// TIA Portal project "SMSS-ENLAB-01-003-1508-012-PLC-B_V13_SP1_1_V17" (V17)

(* hardware
DEVICE "SIMATIC 1200 station_1"  S71200.Device
   slot 0: "S7-1200 rack"  Rack  V1.0
   slot 1: "S7-1200"  CPU 1214C DC/DC/DC  6ES7 214-1AG40-0XB0  V4.5
   slot 2: "DI16 x 24VDC_1"  6ES7 221-1BH30-0XB0  V1.0
   slot 3: "DI8 x 24VDC_1"  6ES7 221-1BF30-0XB0  V1.0
   slot 4: "DQ16 x 24VDC_1"  6ES7 222-1BH30-0XB0  V1.0
DEVICE "HMI"  KTP600 Basic mono PN
   slot 0: "HMI"  HMI  6AV6 647-0AB11-3AX0  12.0.0.0
   slot 1: "HMI_RT_1"  KTP600 Basic mono PN  6AV6 647-0AB11-3AX0  12.0.0.0
   slot 5: "IE_CP_1"  PROFINET Interface  IE_CP  V7.1.0
      slot 1: "PROFINET_Interface_1"  PROFINET Interface
         slot 1: "PORT_1"  Port  1.0.0.0
DEVICE "ET 200S station_1"  ET 200S station
   slot 0: "Rack"  Rail
   slot 0: "IO device_1"  IM 151-3 PN ST  6ES7 151-3AA23-0AB0  V7.0
   slot 1: "PM-E 24VDC_1"  PM-E 24VDC  6ES7 138-4CA01-0AA0
   slot 2: "8DI x 24VDC_1"  8DI DC24V  6ES7 131-4BF00-0AA0
   slot 3: "8DI x 24VDC / SRC ST_1"  8DI DC24V/SRC ST  6ES7 131-4BF50-0AA0
   slot 4: "8DO x 24VDC / 0.5A_1"  8DO DC24V/0.5A  6ES7 132-4BF00-0AA0
DEVICE "CSM"  SCALANCE X-Station
   slot 0: "SCALANCE X rack"  Rail
   slot 0: "CSM 1277 Simatic Net"  6GK7 277-1AA10-0AA0  V1.0
*)

// ===== PLC "S7-1200"  CPU 1214C DC/DC/DC =====

VAR_GLOBAL   // PLC tag table "Default tag table"
   "Flag Negatif Imaje Not ready" AT %M500.2 : Bool;
   "RSAddReject1" AT %I5.5 : Bool;
   "Flag Modu Motor" AT %M300.0 : Bool;
   "RSAddReject2" AT %I5.6 : Bool;
   "PneuAddReject2" AT %Q4.7 : Bool;
   "PSAddReject3" AT %I6.7 : Bool;
   "Reject Conveyor Out" AT %M217.3 : Bool;
   "FP_Reject Conveyor" AT %M219.0 : Bool;
   "Flag P Bad Read" AT %M219.1 : Bool;
   "Error Input Full" AT %M219.2 : Bool;
   "Photosensor 11 Fast Moving" AT %I2.6 : Bool;
   "Always Bad Read Sloft" AT %M217.4 : Bool;
   "Reset Counter Always Bad Read" AT %M217.2 : Bool;
   "FN Imaje 1" AT %M217.5 : Bool;
   "Kosong" AT %I1.4 : Bool;
   "Emergency Stop Push" AT %I4.7 : Bool;
   "Tag_1" AT %I1.0 : Bool;
   "Tag_2" AT %I1.1 : Bool;
   "Tag_3" AT %I0.0 : Bool;
   "Tag_4" AT %Q0.0 : Bool;
   "Tag_5" AT %Q0.1 : Bool;
   "RS_Bypass_Addrej" AT %M31.4 : Bool;
   "PSAddReject1" AT %I5.7 : Bool;
END_VAR

VAR_GLOBAL   // PLC tag table "Output"
   "Reset Error" AT %Q0.4 : Bool;   // Reset Error
   "Pneumatic 1" AT %Q2.0 : Bool;   // Press Heater
   "Pneumatic 2" AT %Q2.1 : Bool;   // Pneumatic Queue
   "Pneumatic 3" AT %Q2.2 : Bool;   // Pneumatic Stopper Label
   "Pneumatic 4" AT %Q2.3 : Bool;   // Pneumatic Stopper Rejector
   "Pneumatic 5" AT %Q2.4 : Bool;   // Pneumatic Rejector
   "Imaje Output Start" AT %Q2.6 : Bool;   // Start Button Markem
   "Imaje Output Pause" AT %Q2.7 : Bool;   // Pause Markem
   "Imaje Output Trigger" AT %Q3.0 : Bool;   // Trigger Markem
   "Red Light" AT %Q3.3 : Bool;   // Red Tower Light
   "Yellow Light" AT %Q3.4 : Bool;   // Yellow Tower Light
   "Green Light" AT %Q3.5 : Bool;   // Green Tower Light
   "Barcode Output PNP" AT %Q1.0 : Bool;   // Output Trigger Barcode
   "Error Output" AT %Q1.1 : Bool;   // Error Output Untuk Digabungkan dengan mesin lain
   "Trigger Mesin Sebelumnya" AT %Q3.1 : Bool;   // Trigger Mesin Pendorong
   "Motor" AT %Q3.6 : Bool;   // Motor Conveyor
   "Teach In Barcode" AT %Q0.5 : Bool;   // Scan and Save Barcode
   "Kran Angin" AT %Q0.6 : Bool;   // Switch Air Valve
   "Pneumatic Pusher" AT %Q4.0 : Bool;
   "Pneumatic Stopper 3 Way" AT %Q4.1 : Bool;
   "Motor Conveyor Pusher" AT %Q4.2 : Bool;
   "PneuAddReject1" AT %Q4.3 : Bool;
   "Red Light FC" AT %Q4.4 : Bool;
   "Yellow Light FC" AT %Q4.5 : Bool;
   "Green Light FC" AT %Q4.6 : Bool;
   "Buzzer AC" AT %Q3.2 : Bool;
END_VAR

VAR_GLOBAL   // PLC tag table "Input"
   "Photosensor 1" AT %I2.0 : Bool;   // Sebelum masuk Heating Tunnel
   "Photosensor 2" AT %I2.1 : Bool;   // Melihat barang batas buffer terakhir
   "Photosensor 11 Fast Moving2" AT %I2.2 : Bool;   // Melihat barang pada slof keluar
   "Photosensor 4" AT %I2.3 : Bool;   // Melihat barang pada tempat label
   "Photosensor 5" AT %I2.4 : Bool;   // Melihat barang pada tempat rejector
   "Reed Switch 1 Advance" AT %I5.0 : Bool;   // Reed Switch Pneumatic 1 Maju
   "Reed Switch 3 Up" AT %I0.2 : Bool;   // Reed Switch Pneumatic 3 Up
   "Reed Switch 3 Down" AT %I0.3 : Bool;   // Reed Switch Pneumatic 3 Down
   "Reed Switch 4 Down" AT %I0.4 : Bool;   // Reed Switch Pneumatic 4 Down
   "Reed Switch 4 Up" AT %I0.5 : Bool;   // Reed Switch Pneumatic 4 Up
   "Reed Switch 5 Advance" AT %I0.6 : Bool;   // Reed Switch Pneumatic 5 Maju
   "Reed Switch 5 Retract" AT %I0.7 : Bool;   // Reed Switch Pneumatic 5 Mundur
   "Imaje 1" AT %I3.0 : Bool;   // Imaje Status Available
   "Imaje 2" AT %I3.1 : Bool;   // Imaje Status Ready
   "Imaje 3" AT %I3.2 : Bool;   // Imaje Status Aplicator Busy (Markem Jalan)
   "Imaje 4" AT %I3.3 : Bool;   // Imaje Status Paper / Ribbon Out
   "Imaje 5" AT %I3.4 : Bool;   // Imaje Status System Error
   "Door Open" AT %I4.3 : Bool;   // Door Open Available
   "PB Run" AT %I4.0 : Bool;   // Push Button Run
   "PB Stop" AT %I4.1 : Bool;   // Push Button Stop
   "PB Reset Error" AT %I4.2 : Bool;   // Push Button Reset Error
   "Pressure Regulator" AT %I1.5 : Bool;   // Mengetahui Tekanan Angin
   "Proximity Markem" AT %I2.7 : Bool;   // Proximity Sensor Untuk Lihat Markem Dibuka
   "PB Machine Bypass" AT %I3.5 : Bool;   // Button Bypass Machine
   "Photosensor 6" AT %I6.0 : Bool;   // Slof Ready on Pusher
   "Photosensor 7" AT %I6.1 : Bool;   // Chute Heating Roll
   "Photosensor 8" AT %I6.2 : Bool;   // Chute 3Way
   "Photosensor 9" AT %I6.3 : Bool;   // Manual Slof Focke
   "PB Run FC" AT %I5.2 : Bool;   // Push Button Run Focke Chute
   "PB Stop FC" AT %I5.3 : Bool;   // Push Button Stop Focke Chute
   "PB Reset Error FC" AT %I5.4 : Bool;   // Push Button Reset Error Focke Chute
   "Door Open FC" AT %I6.5 : Bool;   // Door Open Focke Chute
   "PSAddReject2" AT %I6.6 : Bool;
   "Proximity 10" AT %I6.4 : Bool;   // Door Open FC
   "Reed Switch 1 Retract" AT %I5.1 : Bool;
   "Good Read Barcode" AT %I3.6 : Bool;   // Scanning Goodread
   "Bad Read Barcode" AT %I3.7 : Bool;   // Scanning Badread
   "Photosensor 10" AT %I4.4 : Bool;
END_VAR

VAR_GLOBAL   // PLC tag table "Test Mode"
   "PB Test Mode" AT %M205.0 : Bool;   // PB Test Mode HMI
   "PB Test Pneumatic 1" AT %M205.1 : Bool;
   "PB Test Pneumatic 2" AT %M205.2 : Bool;
   "PB Test Pneumatic 3" AT %M205.3 : Bool;
   "PB Test Pneumatic 4" AT %M205.4 : Bool;
   "PB Test Pneumatic 5" AT %M205.5 : Bool;
   "PB Test Manual Servo" AT %M205.6 : Bool;
   "PB Test Motor" AT %M205.7 : Bool;
   "PB Test Imaje" AT %M206.0 : Bool;
   "PB Test Air Valve" AT %M206.1 : Bool;
   "PB Test Conveyor" AT %M206.3 : Bool;
   "PB Test Pneumatic 6" AT %M206.2 : Bool;
   "PB Test Motor Coveyor Pusher" AT %M206.4 : Bool;
   "PB Test Motor Heating Roll" AT %M206.5 : Bool;
END_VAR

VAR_GLOBAL   // PLC tag table "Flag Output"
   "Flag Direction Servo 1" AT %M210.0 : Bool;
   "Flag Red Light" AT %M210.2 : Bool;
   "Flag Yellow Light" AT %M210.3 : Bool;
   "Flag Green Light" AT %M210.4 : Bool;
   "Flag Pneumatic 1" AT %M211.0 : Bool;
   "Flag Pneumatic 2" AT %M211.1 : Bool;
   "Flag Pneumatic 3" AT %M211.2 : Bool;
   "Flag Pneumatic 4" AT %M211.3 : Bool;
   "Flag Pneumatic 5" AT %M211.4 : Bool;
   "Flag Motor" AT %M211.5 : Bool;
   "Flag Reset Error" AT %M210.6 : Bool;   // Reset Error HMI
   "Flag Direction Servo 2" AT %M210.1 : Bool;
   "Flag Barcode Output" AT %M210.5 : Bool;
   "Flag Imaje Start" AT %M212.0 : Bool;
   "Flag Imaje Pause" AT %M212.1 : Bool;
   "Flag Imaje Trigger" AT %M212.2 : Bool;
   "Flag Mesin Sebelumnya" AT %M212.3 : Bool;
   "Flag Teach In Barcode" AT %M212.4 : Bool;
   "Flag Kran Angin" AT %M212.5 : Bool;
   "Flag Pneumatic 6" AT %M211.6 : Bool;
   "Flag Conveyor" AT %M211.7 : Bool;
   "Flag Motor Conveyor Pusher" AT %M212.6 : Bool;
   "Flag Motor Heating Roll" AT %M212.7 : Bool;
END_VAR

VAR_GLOBAL   // PLC tag table "Cek Pneumatic"
   "Set Flag Cek Pneumatic 1 Maju Bagian Atas" AT %M220.0 : Bool;
   "Set Flag Cek Pneumatic 1 Maju Bagian Bawah" AT %M220.1 : Bool;
   "Flag RS Pneumatic 1 Pusher  Advance" AT %M220.2 : Bool;
   "Flag RS Pneumatic 1 Retract" AT %M220.3 : Bool;
   "Flag RS Pneumatic 1 Advance Error" AT %M220.4 : Bool;
   "Flag RS Pneumatic 1 Retract Error" AT %M220.5 : Bool;
   "Set Flag Cek Pneumatic 3 Maju" AT %M221.0 : Bool;
   "Set Flag Cek Pneumatic 3 Mundur" AT %M221.1 : Bool;
   "Flag RS Pneumatic 3 Up" AT %M221.2 : Bool;
   "Flag  RS Pneumatic 3 Down" AT %M221.3 : Bool;
   "Flag RS Pneumatic 3 Up Error" AT %M221.4 : Bool;
   "Flag RS Pneumatic 3 Down Error" AT %M221.5 : Bool;
   "Set Flag Cek Pneumatic 4 Maju" AT %M222.0 : Bool;
   "Set Flag Cek Pneumatic 4 Mundur" AT %M222.1 : Bool;
   "Flag RS Pneumatic 4 Down" AT %M222.2 : Bool;
   "Flag RS Pneumatic 4 Up" AT %M222.3 : Bool;
   "Flag RS Pneumatic 4 Down Error" AT %M222.4 : Bool;
   "Flag RS Pneumatic 4 Up Error" AT %M222.5 : Bool;
   "Set Flag Cek Pneumatic 5 Maju" AT %M223.0 : Bool;
   "Set Flag Cek Pneumatic 5 Mundur" AT %M223.1 : Bool;
   "Flag RS Pneumatic 5 Advance" AT %M223.2 : Bool;
   "Flag RS Pneumatic 5 Retract" AT %M223.3 : Bool;
   "Flag RS Pneumatic 5 Advnance Error" AT %M223.4 : Bool;
   "Flag RS Pneumatic 5 Retract Error" AT %M223.5 : Bool;
END_VAR

VAR_GLOBAL   // PLC tag table "Flag Machine"
   "Machine Running" AT %M200.0 : Bool;
   "Flag Stop" AT %M200.3 : Bool;
   "Block 2 Ready" AT %M230.0 : Bool;
   "Flag Good Read Barcode" AT %M230.1 : Bool;
   "Flag Bad Read Barcode" AT %M230.2 : Bool;
   "Flag Ejector Jalan" AT %M230.3 : Bool;
   "Slof Ready" AT %M230.4 : Bool;
   "Flag Stamp Finish" AT %M230.5 : Bool;
   "Enable Barcode" AT %M230.6 : Bool;
   "Flag Slof Ready" AT %M230.7 : Bool;
   "Flag Sudah Di Datecode" AT %M231.0 : Bool;
   "Flag Sudah Di Barcode" AT %M231.1 : Bool;
   "Flag Good Read Barcode Finish" AT %M231.2 : Bool;
   "Flag Rejector Start" AT %M231.4 : Bool;
   "Flag Barang Sudah Dibuang" AT %M231.5 : Bool;
   "Flag Ready to Reject" AT %M231.6 : Bool;
   "Enable Press Heater" AT %M231.3 : Bool;
   "Flag Heating Ready" AT %M232.0 : Bool;
   "Slof Manual Ready" AT %M232.1 : Bool;
   "Flag Enable/Disable Barcode HMI" AT %M30.0 : Bool;
   "Flag Enable/Disable Error Chute 3 Way" AT %M30.1 : Bool;
   "Disable Barcode" AT %M232.4 : Bool;
   "Disable Heater" AT %M232.5 : Bool;
   "Flag Parameter Page" AT %M232.6 : Bool;
   "Flag Main Page" AT %M232.7 : Bool;
   "Flag Error boleh jalan" AT %M233.0 : Bool;
   "Flag Rejector Finish" AT %M233.1 : Bool;
   "Flag Heater Error HMI" AT %M30.2 : Bool;
   "Flag Reed Switch Bypass" AT %M30.3 : Bool;
   "Flag Machine Bypass" AT %M30.7 : Bool;
   "Flag Enable/Disable Error Chute Before Heating Roll" AT %M30.4 : Bool;
   "Flag Enable/Disable Error Door Open" AT %M30.5 : Bool;
   "Flag Enable/Disable Block Focke" AT %M30.6 : Bool;
   "Flag Ready to Stamp" AT %M233.2 : Bool;
   "Flag Negatif Photosensor 4" AT %M232.3 : Bool;
   "Section Reject" AT %M232.2 : Bool;
   "RS Bypass Pneumatic 1" AT %M31.0 : Bool;
   "RS Bypass Pneumatic 3" AT %M31.1 : Bool;
   "RS Bypass Pneumatic 4" AT %M31.2 : Bool;
   "RS Bypass Pneumatic 5" AT %M31.3 : Bool;
   "Flag Enable/Disable Flow to Reject" AT %M31.5 : Bool;
   "Flag Slof Jamed" AT %M233.3 : Bool;
   "Flow to Reject" AT %M233.4 : Bool;
   "Flag Stopper Heating Finish" AT %M233.5 : Bool;
   "Slof Manual Finish" AT %M234.0 : Bool;
   "Flag Enable/Disable Heating Roll" AT %M31.6 : Bool;
   "Flag Enable/Disable Reject Outfeed" AT %M31.7 : Bool;
   "Flag Buzzer AC" AT %M500.1 : Bool;
   "Flag Negatif Conveyor Outfeed" AT %M500.0 : Bool;
   "Conveyor Outfeed Finish" AT %M216.7 : Bool;
   "Confeyor Outfeed" AT %M217.0 : Bool;
END_VAR

VAR_GLOBAL   // PLC tag table "Counter"
   "Counter" AT %MW5 : Int;
   "Counter PV" AT %MW7 : Int;
   "Reset Counter" AT %M200.1 : Bool;
   "Counter Ejector" AT %MW9 : Int;
   "Previous Scan Sensor Ejector" AT %M200.4 : Bool;
   "Counter PV Ejector" AT %MW11 : Int;
END_VAR

VAR_GLOBAL   // PLC tag table "Timer"
   "Timer Delay Stamp" AT %MD32 : Time;
   "Timer Trigger Barcode" AT %MD39 : Time;
   "Timer Rejector Slof" AT %MD43 : Time;
   "Timer AutoReject" AT %MD48 : Time;
END_VAR

VAR_GLOBAL   // PLC tag table "Flag Error"
   "Error" AT %M215.0 : Bool;   // Flag Error
   "Error Pressure" AT %M215.1 : Bool;
   "Error Door Open" AT %M215.2 : Bool;
   "Error Servo 1" AT %M215.3 : Bool;
   "Error Servo 2" AT %M215.4 : Bool;
   "Servo 1 Not Ready" AT %M215.5 : Bool;
   "Servo 2 Not Ready" AT %M215.6 : Bool;
   "Error Imaje Paper / Ribbon Out" AT %M215.7 : Bool;
   "Error Imaje System" AT %M216.0 : Bool;
   "Markem Not In Position" AT %M216.1 : Bool;
   "Heater Not Ready" AT %M216.2 : Bool;
   "Error Group" AT %MW4 : Word;
   "Markem Not Ready" AT %M216.4 : Bool;
   "Error Door Open FC" AT %M216.5 : Bool;
   "Chute Before Heating Roll Full" AT %M231.7 : Bool;
   "Chute 3 Way Full" AT %M234.1 : Bool;
   "Error Door Open Proximity" AT %M216.3 : Bool;
   "Error Conveyor Outfeed" AT %M217.1 : Bool;
END_VAR

DATA_BLOCK "DB Test Mode"   // DB1
{ S7_Optimized_Access := 'TRUE' }
VERSION : 0.1
// stored: InstanceOfName Block Test Mode
"Block Test Mode"
BEGIN
END_DATA_BLOCK

DATA_BLOCK "DB Error Mode"   // DB2
{ S7_Optimized_Access := 'TRUE' }
VERSION : 0.1
// stored: InstanceOfName Block Error Mode
"Block Error Mode"
BEGIN
END_DATA_BLOCK

DATA_BLOCK "DB Flag Output"   // DB3
{ S7_Optimized_Access := 'TRUE' }
VERSION : 0.1
// stored: InstanceOfName Block Output
"Block Output"
BEGIN
END_DATA_BLOCK

DATA_BLOCK "DB Block Labelling"   // DB25
{ S7_Optimized_Access := 'TRUE' }
VERSION : 0.1
// stored: InstanceOfName Block Labeling
"Block Labeling"
BEGIN
END_DATA_BLOCK

DATA_BLOCK "Data_DTL1"   // DB29
{ S7_Optimized_Access := 'TRUE' }
VERSION : 0.1
   VAR RETAIN
      Input : DTL := DTL#2014-01-01-00:00:00;
      Output : DTL := DTL#2014-01-01-00:00:00;
      Cur_ShiftA : DTL := DTL#1970-01-01-00:00:00;   // Data Awal Shift Yang ngitung terus
      Cur_ShiftA_1 : DTL;
      Cur_ShiftA_2 : DTL;
      Cur_ShiftA_3 : DTL;
      Cur_ShiftA_4 : DTL;
      Cur_ShiftA_5 : DTL;
      Cur_ShiftB : DTL;
      Cur_ShiftB_1 : DTL;
      Cur_ShiftB_2 : DTL;
      Cur_ShiftB_3 : DTL;
      Cur_ShiftB_4 : DTL;
      Cur_ShiftB_5 : DTL;
   END_VAR
BEGIN
END_DATA_BLOCK

DATA_BLOCK "DB Block Focke"   // DB34
{ S7_Optimized_Access := 'TRUE' }
VERSION : 0.1
// stored: InstanceOfName Block Focke
"Block Focke"
BEGIN
END_DATA_BLOCK

DATA_BLOCK "Data_Time"   // DB35
{ S7_Optimized_Access := 'TRUE' }
VERSION : 0.1
   VAR RETAIN
      "Shift 1A" : Time := T#6h;   // Awal Shift Static Sesuai pengaturan
      "Shift 1B" : Time := T#14h;
      "Shift 2A" : Time := T#14h;
      "Shift 2B" : Time := T#22h;
      "Shift 3A" : Time := T#22h;
      "Shift 3B" : Time := T#6h;
      "Shift 1B_Min5" : Time;   // 5 Detik Sebelum Akhir Shift
      "Shift 2B_Min5" : Time;   // 5 Detik Sebelum Akhir Shift
      "Shift 3B_Min5" : Time;   // 5 Detik Sebelum Akhir Shift
      "TOD Sistem" : Time_Of_Day;
      "Time Sistem" : Time;
      "Time Total 1 Shift" : Time;   // Selisih Waktu dalam satu shift/waktu yang di gunakan
      "Timer Delay Stamp" : Time;
      "Timer Trigger Barcode" : Time := T#300ms;
      "Timer Rejector Slof" : Time;
      "Timer AutoReject" : Time := T#300ms;
   END_VAR
BEGIN
END_DATA_BLOCK

DATA_BLOCK "Data_String"   // DB36
{ S7_Optimized_Access := 'TRUE' }
VERSION : 0.1
   VAR RETAIN
      "sDT_Machine id" : String := 'LU 12';
   END_VAR
BEGIN
END_DATA_BLOCK

DATA_BLOCK "Error Alarm"   // DB39
{ S7_Optimized_Access := 'FALSE' }
VERSION : 0.1
   VAR
      "Pressure Low" : Bool;
      "Door Open Labelling" : Bool;
      "Door Open Focke Chute" : Bool;
      "Chute 3Way Full" : Bool;
      "Door Open Proximity" : Bool;
      Static_4 : Bool;
      "Imaje Paper/Ribbon Out" : Bool;
      "Imaje System Error" : Bool;
      "Imaje Not In Position" : Bool;
      "Heater Not Ready" : Bool;
      "Reed Switch Pneumatic 1 Pusher Advance" : Bool;
      "Reed Switch Pneumatic 1 Pusher Retract" : Bool;
      "Reed Switch Pneumatic 3 Up" : Bool;
      "Reed Switch Pneumatic 3 Down" : Bool;
      "Infeed Chute full" : Bool;
   END_VAR
BEGIN
END_DATA_BLOCK

DATA_BLOCK "Error Alarm 2"   // DB40
{ S7_Optimized_Access := 'FALSE' }
VERSION : 0.1
   VAR
      "Reed Switch Pneumatic 4 Down" : Bool;
      "Reed Switch Pneumatic 4 Up" : Bool;
      "Reed Switch Pneumatic 5 Advance" : Bool;
      "Reed Switch Pneumatic 5 Retract" : Bool;
      "Conveyor Outfeed jammed" : Bool;
      "Sloft Jammed In Labelling" : Bool;
      "Slof Jammed Infeed Chute" : Bool;
      "Always Bad Read Sloft" : Bool;
      "Paper Or Ribbon Low" : Bool;
      "Emergency Stop Push" : Bool;
   END_VAR
BEGIN
END_DATA_BLOCK

DATA_BLOCK "Data_Integer"   // DB43
{ S7_Optimized_Access := 'TRUE' }
VERSION : 0.1
   VAR RETAIN
      RV1 : Word;   // RV Baca Date Time
      RV2 : Word;   // RV Set Date Time
      IDay : USInt := 1;
      IMonth : USInt := 1;
      IYear : UInt := 2014;
      IHour : USInt;
      IMinute : USInt;
      ISecond : USInt;
      S1AHour : USInt := 6;
      S1AMinute : USInt;
      S1ASecond : USInt;
      S1BHour : USInt := 14;
      S1BMinute : USInt;
      S1BSecond : USInt;
      S2AHour : USInt := 14;
      S2AMinute : USInt;
      S2ASecond : USInt;
      S2BHour : USInt := 22;
      S2BMinute : USInt;
      S2BSecond : USInt;
      S3AHour : USInt := 22;
      S3AMinute : USInt;
      S3ASecond : USInt;
      S3BHour : USInt := 6;
      S3BMinute : USInt;
      S3BSecond : USInt;
      T_Shift1A : UDInt;
      T_Shift1B : UDInt;
      T_Shift2A : UDInt;
      T_Shift2B : UDInt;
      T_Shift3A : UDInt;
      T_Shift3B : UDInt;
   END_VAR
BEGIN
END_DATA_BLOCK

DATA_BLOCK "Data_Bool1"   // DB44
{ S7_Optimized_Access := 'TRUE' }
VERSION : 0.1
   VAR
      "F_Set Time Day" : Bool;   // Off : Baca date Time Sistem Enable ; On : Eksekusi setting date time sistem
      "F_Set Time Shift" : Bool;
      "FP_In Sloft" : Bool;
      FP_GRead : Bool;
      "FP_GRead Rej" : Bool;
   END_VAR
   VAR RETAIN
      "FP_Flag Shift1" : Bool;
      "FP_Flag Shift2" : Bool;
      "FP_Flag Shift3" : Bool;
      "Flag After Copi 5" : Bool;
      "Flag After Copi 4" : Bool;
      "Flag After Copi 3" : Bool;
      "Flag After Copi 2" : Bool;
      "Flag After Copi 1" : Bool;
      "Flag AfterHapus Data" : Bool;
   END_VAR
   VAR
      "FN_Hapus data" : Bool;
      "Flag Hapus Data" : Bool;
      "FPN_Hitung Frek Error" : Array[1..15] of Bool;
      "Flag After Hitung Frek Error" : Array[1..7] of Bool;
   END_VAR
   VAR RETAIN
      "Flag Copy Data" : Bool;
      "Flag Copy Data_2" : Bool;
      "Flag Shift 1" : Bool;
      "Flag Shift 2" : Bool;
      "Flag Shift 3" : Bool;
   END_VAR
   VAR
      "Flag_Cek Shift" : Array[1..3] of Bool;
   END_VAR
   VAR RETAIN
      "Stop Baca" : Bool;
   END_VAR
BEGIN
END_DATA_BLOCK

DATA_BLOCK "AddReject2_DB"   // DB46
{ S7_Optimized_Access := 'TRUE' }
VERSION : 0.1
// stored: InstanceOfName AddReject2
"AddReject2"
BEGIN
END_DATA_BLOCK

DATA_BLOCK "Data_TimeData"   // DB50
{ S7_Optimized_Access := 'TRUE' }
VERSION : 0.1
   VAR RETAIN
      "T_Imaje Er" : Time;
      "T_Imaje Er_A" : Time;
      "T_Imaje Er_B" : Time;
      "T_Slof Jam1" : Time;
      "T_Slof Jam1_A" : Time;
      "T_Slof Jam1_B" : Time;
      "T_Down Stop" : Time;
      "T_Down Stop_A" : Time;
      "T_Down Stop_B" : Time;
      "T_RS Pneu Er" : Time;
      "T_RS Pneu Er_A" : Time;
      "T_RS Pneu Er_B" : Time;
      "T_Paper R Out" : Array[0..2] of Time;
      "T_Imaje Not In Position" : Array[0..2] of Time;
      "Mesin Run" : Time;
      "Mesin Run_A" : Time;
      "Mesin Run_B" : Time;
      "Mesin Run Baypass" : Time;
      "Mesin Run Baypass_A" : Time;
      "Mesin Run Baypass_B" : Time;
      "Mesin Stop" : Time;
      "Mesin Stop_A" : Time;
      "Mesin Stop_B" : Time;
      "Mesin Error" : Time;
      "Mesin Error_A" : Time;
      "Mesin Error_B" : Time;
      "Total Time Machine" : Time;
      "T_Always bad Read" : Time;
   END_VAR
   VAR
      "T_Always bad Read_A" : Time;
      "T_Always bad Read_B" : Time;
   END_VAR
   VAR RETAIN
      "T_Press Low" : Time;
   END_VAR
   VAR
      "T_Press Low_A" : Time;
      "T_Press Low_B" : Time;
   END_VAR
   VAR RETAIN
      "T_Door Open" : Time;
   END_VAR
   VAR
      "T_Door Open_A" : Time;
      "T_Door Open_B" : Time;
   END_VAR
   VAR RETAIN
      "T_Total Detail Error" : Time;
   END_VAR
BEGIN
END_DATA_BLOCK

DATA_BLOCK "Data_Real"   // DB51
{ S7_Optimized_Access := 'TRUE' }
VERSION : 0.1
   VAR RETAIN
      "R  Good R" : Real;
      "R Bad Read" : Real;
      "R Input Sloft" : Real;
      "R Reject Out Stop" : Real;
      "R Total Output" : Real;
      "Sloft Bypass" : Real;
      InputReject : Real;
      "%Bad Read" : Array[0..5] of Real;
      "%Good Read" : Array[0..5] of Real;
      "% Reject Out Stop" : Array[0..5] of Real;
      "%InputReject" : Array[0..5] of Real;
      "% label Sloft" : Array[0..5] of Real;
      "% Unlabel Sloft" : Array[0..5] of Real;
      "% Sloft bypass" : Array[0..5] of Real;
      "% Total Output" : Array[0..5] of Real;
      "R Total 1 Shift" : Real;
      "R Mesin Run" : Real;
      "R Mesin Run Baypass" : Real;
      "R Mesin Stop" : Real;
      "R Mesin error" : Real;
      "R Downstream stop" : Real;
      "%Mesin Run" : Array[0..5] of Real;
      "%Mesin Run Baypass" : Array[0..5] of Real;
      "%Mesin Stop" : Array[0..5] of Real;
      "%Mesin Error" : Array[0..5] of Real;
      "%Downstream stop" : Array[0..5] of Real;
   END_VAR
BEGIN
END_DATA_BLOCK

DATA_BLOCK "Data_IntData"   // DB53
{ S7_Optimized_Access := 'TRUE' }
VERSION : 0.1
   VAR RETAIN
      "Good R" : UDInt;
      "Good R_1" : UDInt := 0;
      "Good R_2" : UDInt := 0;
      "Good R_3" : UDInt := 0;
      "Good R_4" : UDInt := 0;
      "Good R_5" : UDInt := 0;
      "Reject Out S" : UDInt;
      "Reject Out S_1" : UDInt := 0;
      "Reject Out S_2" : UDInt := 0;
      "Reject Out S_3" : UDInt := 0;
      "Reject Out S_4" : UDInt := 0;
      "Reject Out S_5" : UDInt := 0;
      "Bad R" : UDInt;
      "Bad R_1" : UDInt := 0;
      "Bad R_2" : UDInt := 0;
      "Bad R_3" : UDInt := 0;
      "Bad R_4" : UDInt := 0;
      "Bad R_5" : UDInt;
      InReject : UDInt;
      InReject_1 : UDInt;
      InReject_2 : UDInt;
      InReject_3 : UDInt;
      InReject_4 : UDInt;
      InReject_5 : UDInt;
      "Sloft Bypass" : Array[0..5] of UDInt;
      "Label Sloft" : Array[0..5] of UDInt;
      "Un label Sloft" : Array[0..5] of UDInt;
      "Tot Out Slof" : UDInt;
      "Tot Out Slof_1" : UDInt;
      "Tot Out Slof_2" : UDInt;
      "Tot Out Slof_3" : UDInt;
      "Tot Out Slof_4" : UDInt;
      "Tot Out Slof_5" : UDInt;
      "Input Sloft" : UDInt;   // Data Input Sloft
      "Input Sloft_1" : UDInt := 0;
      "Input Sloft_2" : UDInt := 0;
      "Input Sloft_3" : UDInt := 0;
      "Input Sloft_4" : UDInt := 0;
      "Input Sloft_5" : UDInt := 0;
      "Int Mesin Run" : UDInt;
      "Int Mesin Run Baypass" : UDInt;
      "Int Mesin Stop" : UDInt;
      "Int Mesin error" : UDInt;
      "Int Downstream stop" : UDInt;
      "uintDT_Imaje Trigger" : Array[0..5] of UInt;
      "uintDT_Imaje Busy" : Array[0..5] of UInt;
      uintDT_AplicatorFreeze : Array[0..5] of UInt;
   END_VAR
BEGIN
END_DATA_BLOCK

DATA_BLOCK "Data_integer2"   // DB54
{ S7_Optimized_Access := 'TRUE' }
VERSION : 0.1
   VAR RETAIN
      T_Shift1B_Min5 : UDInt;   // 5 Detik sebelum akhir Shift 1
      T_Shift2B_Min5 : UDInt;   // 5 Detik sebelum akhir Shift 1
      T_Shift3B_Min5 : UDInt;   // 5 Detik sebelum akhir Shift 1
      "Flag Power Off" : USInt := 1;   // Harus Di Isi Pas Mulai Download sesuai sama shiftnya
      "Flag Input Always Bad Read" : USInt := 5;
      "Int Total 1 Shift" : UDInt;
   END_VAR
BEGIN
END_DATA_BLOCK

DATA_BLOCK "S Block Par Statistika_DB"   // DB56
{ S7_Optimized_Access := 'TRUE' }
VERSION : 0.1
// stored: InstanceOfName S Block Par Statistika
"S Block Par Statistika"
BEGIN
END_DATA_BLOCK

DATA_BLOCK "S Check Range Shift_DB"   // DB57
{ S7_Optimized_Access := 'TRUE' }
VERSION : 0.1
// stored: InstanceOfName S Check Range Shift
"S Check Range Shift"
BEGIN
END_DATA_BLOCK

DATA_BLOCK "S Block Current Shift_DB"   // DB58
{ S7_Optimized_Access := 'TRUE' }
VERSION : 0.1
// stored: InstanceOfName S Block Current Shift
"S Block Current Shift"
BEGIN
END_DATA_BLOCK

DATA_BLOCK "S Block Current Shift_M5_DB"   // DB59
{ S7_Optimized_Access := 'TRUE' }
VERSION : 0.1
// stored: InstanceOfName S Block Current Shift_M5
"S Block Current Shift_M5"
BEGIN
END_DATA_BLOCK

DATA_BLOCK "S Block Current Shift_M4_DB"   // DB61
{ S7_Optimized_Access := 'TRUE' }
VERSION : 0.1
// stored: InstanceOfName S Block Current Shift_M4
"S Block Current Shift_M4"
BEGIN
END_DATA_BLOCK

DATA_BLOCK "S Block Current Shift_M3_DB"   // DB62
{ S7_Optimized_Access := 'TRUE' }
VERSION : 0.1
// stored: InstanceOfName S Block Current Shift_M3
"S Block Current Shift_M3"
BEGIN
END_DATA_BLOCK

DATA_BLOCK "S Block Current Shift_M2_DB"   // DB63
{ S7_Optimized_Access := 'TRUE' }
VERSION : 0.1
// stored: InstanceOfName S Block Current Shift_M2
"S Block Current Shift_M2"
BEGIN
END_DATA_BLOCK

DATA_BLOCK "S Block Current Shift_M1_DB"   // DB64
{ S7_Optimized_Access := 'TRUE' }
VERSION : 0.1
// stored: InstanceOfName S Block Current Shift_M1
"S Block Current Shift_M1"
BEGIN
END_DATA_BLOCK

DATA_BLOCK "Data_DTLData"   // DB66
{ S7_Optimized_Access := 'TRUE' }
VERSION : 0.1
   VAR RETAIN
      "DTL_Imaje Er" : DTL;
      "DTL_Imaje Er_1" : DTL;
      "DTL_Imaje Er_2" : DTL;
      "DTL_Imaje Er_3" : DTL;
      "DTL_Imaje Er_4" : DTL;
      "DTL_Imaje Er_5" : DTL;
      "DTL_Sloft Jam1" : DTL;
      "DTL_Sloft Jam1_1" : DTL;
      "DTL_Sloft Jam1_2" : DTL;
      "DTL_Sloft Jam1_3" : DTL;
      "DTL_Sloft Jam1_4" : DTL;
      "DTL_Sloft Jam1_5" : DTL;
      "DTL_Down Stop" : DTL;
      "DTL_Down Stop_1" : DTL;
      "DTL_Down Stop_2" : DTL;
      "DTL_Down Stop_3" : DTL;
      "DTL_Down Stop_4" : DTL;
      "DTL_Down Stop_5" : DTL;
      "DTL_RS Pneu Er" : DTL;
      "DTL_RS Pneu Er_1" : DTL;
      "DTL_RS Pneu Er_2" : DTL;
      "DTL_RS Pneu Er_3" : DTL;
      "DTL_RS Pneu Er_4" : DTL;
      "DTL_RS Pneu Er_5" : DTL;
      "DTL_Paper R Out" : Array[0..5] of DTL;
      "DTL_Imaje Not In Position" : Array[0..5] of DTL;
      "DTL_Mesin Run" : Array[0..5] of DTL;
      "DTL_Mesin Run Baypass" : Array[0..5] of DTL;
      "DTL_Mesin Stop" : Array[0..5] of DTL;
      "DTL_Mesin Error" : Array[0..5] of DTL;
      "Total Time Machine" : Array[0..5] of DTL;
      "DTL_Always bad Read" : Array[0..5] of DTL;
      "DTL_Press Low" : Array[0..5] of DTL;
      "DTL_Door Open" : Array[0..5] of DTL;
      "DTL_Total Detail Error" : Array[0..5] of DTL;
   END_VAR
BEGIN
END_DATA_BLOCK

DATA_BLOCK "Data_TODData"   // DB72
{ S7_Optimized_Access := 'TRUE' }
VERSION : 0.1
   VAR RETAIN
      "TOD_Imaje Er" : Time_Of_Day;
      "TOD_Sloft Jam1" : Time_Of_Day;
      "TOD_Down Stop" : Time_Of_Day;
      "TOD_RS Pneu Er" : Time_Of_Day;
      "TOD_Paper R Out" : Time_Of_Day;
      "Imaje Not In Position" : Time_Of_Day;
      "TOD_Cur Static ShiftA" : Array[0..5] of Time_Of_Day;   // Batas Awal currect Shift static
      "TOD_Mesin Run" : Time_Of_Day;
      "TOD_Mesin Run Baypass" : Time_Of_Day;
      "TOD_Mesin Stop" : Time_Of_Day;
      "TOD_Mesin Error" : Time_Of_Day;
      "Total Time Machine" : Time_Of_Day;
      "TOD_Always bad Read" : Time_Of_Day;
   END_VAR
   VAR
      "TOD_Press Low" : Time_Of_Day;
      "TOD_Door Open" : Time_Of_Day;
      "TOD_Total Detail Error" : Time_Of_Day;
   END_VAR
BEGIN
END_DATA_BLOCK

DATA_BLOCK "S Block Hapus Data_DB"   // DB77
{ S7_Optimized_Access := 'TRUE' }
VERSION : 0.1
// stored: InstanceOfName S Block Hapus Data
"S Block Hapus Data"
BEGIN
END_DATA_BLOCK

DATA_BLOCK "Data_Bool2"   // DB89
{ S7_Optimized_Access := 'TRUE' }
VERSION : 0.1
   VAR
      "bFL_Emergency Stop" : Bool;
      "bFL_Error Imaje" : Bool;
      "bFL_FP Flow Reject" : Bool;
      "bFL_Hitung Out Sloft Baypass Mesin" : Bool;
      "bFL_FP Sloft Bypasss" : Bool;
      "bFL_error Imaje Baypass other" : Bool;
      "bFL_Flag Positif Output Trigger" : Bool;
      "bFL_Flag Positif Imaje 3" : Bool;
      "Sloft jam labelling" : Bool;
      "Reset Alarm" : Bool;
      FP_RejInput : Bool;
   END_VAR
BEGIN
END_DATA_BLOCK

// folder: System blocks/Program resources

DATA_BLOCK "Timer Error PS Pneumatic 1 Retract Error"   // DB4
{ S7_Optimized_Access := 'TRUE' }
AUTHOR : Simatic
FAMILY : IEC
NAME : IEC_TMR
VERSION : 1.0
// stored: InstanceOfName IEC_TIMER
"IEC_TIMER"
BEGIN
END_DATA_BLOCK

DATA_BLOCK "ttM_TimerAddRej1"   // DB5
{ S7_Optimized_Access := 'TRUE' }
AUTHOR : Simatic
FAMILY : IEC
NAME : IEC_TMR
VERSION : 1.0
// stored: InstanceOfName IEC_TIMER
"IEC_TIMER"
BEGIN
END_DATA_BLOCK

DATA_BLOCK "Timer PS Pneumatic 1 Advance"   // DB6
{ S7_Optimized_Access := 'TRUE' }
AUTHOR : Simatic
FAMILY : IEC
NAME : IEC_TMR
VERSION : 1.0
// stored: InstanceOfName IEC_TIMER
"IEC_TIMER"
BEGIN
END_DATA_BLOCK

DATA_BLOCK "Timer Error RS Pneumatic 1 Advance Error"   // DB7
{ S7_Optimized_Access := 'TRUE' }
AUTHOR : Simatic
FAMILY : IEC
NAME : IEC_TMR
VERSION : 1.0
// stored: InstanceOfName IEC_TIMER
"IEC_TIMER"
BEGIN
END_DATA_BLOCK

DATA_BLOCK "Timer RS Pneumatic 3 Up Error"   // DB8
{ S7_Optimized_Access := 'TRUE' }
AUTHOR : Simatic
FAMILY : IEC
NAME : IEC_TMR
VERSION : 1.0
// stored: InstanceOfName IEC_TIMER
"IEC_TIMER"
BEGIN
END_DATA_BLOCK

DATA_BLOCK "Timer RS Pneumatic 3 Up"   // DB9
{ S7_Optimized_Access := 'TRUE' }
AUTHOR : Simatic
FAMILY : IEC
NAME : IEC_TMR
VERSION : 1.0
// stored: InstanceOfName IEC_TIMER
"IEC_TIMER"
BEGIN
END_DATA_BLOCK

DATA_BLOCK "Timer RS Pneumatic 3 Down Error"   // DB10
{ S7_Optimized_Access := 'TRUE' }
AUTHOR : Simatic
FAMILY : IEC
NAME : IEC_TMR
VERSION : 1.0
// stored: InstanceOfName IEC_TIMER
"IEC_TIMER"
BEGIN
END_DATA_BLOCK

DATA_BLOCK "Timer RS Pneumatic 3 Down"   // DB11
{ S7_Optimized_Access := 'TRUE' }
AUTHOR : Simatic
FAMILY : IEC
NAME : IEC_TMR
VERSION : 1.0
// stored: InstanceOfName IEC_TIMER
"IEC_TIMER"
BEGIN
END_DATA_BLOCK

DATA_BLOCK "Timer RS Pneumatic 4 Down Error"   // DB12
{ S7_Optimized_Access := 'TRUE' }
AUTHOR : Simatic
FAMILY : IEC
NAME : IEC_TMR
VERSION : 1.0
// stored: InstanceOfName IEC_TIMER
"IEC_TIMER"
BEGIN
END_DATA_BLOCK

DATA_BLOCK "Timer RS Pneumatic 4 Down"   // DB13
{ S7_Optimized_Access := 'TRUE' }
AUTHOR : Simatic
FAMILY : IEC
NAME : IEC_TMR
VERSION : 1.0
// stored: InstanceOfName IEC_TIMER
"IEC_TIMER"
BEGIN
END_DATA_BLOCK

DATA_BLOCK "Timer RS Pneumatic 4 Up Error"   // DB14
{ S7_Optimized_Access := 'TRUE' }
AUTHOR : Simatic
FAMILY : IEC
NAME : IEC_TMR
VERSION : 1.0
// stored: InstanceOfName IEC_TIMER
"IEC_TIMER"
BEGIN
END_DATA_BLOCK

DATA_BLOCK "Timer RS Pneumatic 4 Up"   // DB15
{ S7_Optimized_Access := 'TRUE' }
AUTHOR : Simatic
FAMILY : IEC
NAME : IEC_TMR
VERSION : 1.0
// stored: InstanceOfName IEC_TIMER
"IEC_TIMER"
BEGIN
END_DATA_BLOCK

DATA_BLOCK "Timer RS Pneumatic 5 Advance Error"   // DB16
{ S7_Optimized_Access := 'TRUE' }
AUTHOR : Simatic
FAMILY : IEC
NAME : IEC_TMR
VERSION : 1.0
// stored: InstanceOfName IEC_TIMER
"IEC_TIMER"
BEGIN
END_DATA_BLOCK

DATA_BLOCK "Timer RS Pneumatic 5 Advance"   // DB17
{ S7_Optimized_Access := 'TRUE' }
AUTHOR : Simatic
FAMILY : IEC
NAME : IEC_TMR
VERSION : 1.0
// stored: InstanceOfName IEC_TIMER
"IEC_TIMER"
BEGIN
END_DATA_BLOCK

DATA_BLOCK "Timer RS Pneumatic 5 Retract Error"   // DB18
{ S7_Optimized_Access := 'TRUE' }
AUTHOR : Simatic
FAMILY : IEC
NAME : IEC_TMR
VERSION : 1.0
// stored: InstanceOfName IEC_TIMER
"IEC_TIMER"
BEGIN
END_DATA_BLOCK

DATA_BLOCK "Timer RS Pneumatic 5 Retract"   // DB19
{ S7_Optimized_Access := 'TRUE' }
AUTHOR : Simatic
FAMILY : IEC
NAME : IEC_TMR
VERSION : 1.0
// stored: InstanceOfName IEC_TIMER
"IEC_TIMER"
BEGIN
END_DATA_BLOCK

DATA_BLOCK "Timer Error Chute 3 Way"   // DB20
{ S7_Optimized_Access := 'TRUE' }
AUTHOR : Simatic
FAMILY : IEC
NAME : IEC_TMR
VERSION : 1.0
// stored: InstanceOfName IEC_TIMER
"IEC_TIMER"
BEGIN
END_DATA_BLOCK

DATA_BLOCK "Timer Buzzer AC1"   // DB21
{ S7_Optimized_Access := 'TRUE' }
AUTHOR : Simatic
FAMILY : IEC
NAME : IEC_TMR
VERSION : 1.0
// stored: InstanceOfName IEC_TIMER
"IEC_TIMER"
BEGIN
END_DATA_BLOCK

DATA_BLOCK "Safety Slof jammed"   // DB22
{ S7_Optimized_Access := 'TRUE' }
AUTHOR : Simatic
FAMILY : IEC
NAME : IEC_TMR
VERSION : 1.0
// stored: InstanceOfName IEC_TIMER
"IEC_TIMER"
BEGIN
END_DATA_BLOCK

DATA_BLOCK "Timer Slof Jamed"   // DB23
{ S7_Optimized_Access := 'TRUE' }
AUTHOR : Simatic
FAMILY : IEC
NAME : IEC_TMR
VERSION : 1.0
// stored: InstanceOfName IEC_TIMER
"IEC_TIMER"
BEGIN
END_DATA_BLOCK

DATA_BLOCK "IEC_Timer_Tunggu_Barcode_DB"   // DB24
{ S7_Optimized_Access := 'TRUE' }
AUTHOR : Simatic
FAMILY : IEC
NAME : IEC_TMR
VERSION : 1.0
// stored: InstanceOfName IEC_TIMER
"IEC_TIMER"
BEGIN
END_DATA_BLOCK

DATA_BLOCK "Timer Chute Before Heating Roll"   // DB26
{ S7_Optimized_Access := 'TRUE' }
AUTHOR : Simatic
FAMILY : IEC
NAME : IEC_TMR
VERSION : 1.0
// stored: InstanceOfName IEC_TIMER
"IEC_TIMER"
BEGIN
END_DATA_BLOCK

DATA_BLOCK "IEC_Timer_Stempel_DB"   // DB27
{ S7_Optimized_Access := 'TRUE' }
AUTHOR : Simatic
FAMILY : IEC
NAME : IEC_TMR
VERSION : 1.0
// stored: InstanceOfName IEC_TIMER
"IEC_TIMER"
BEGIN
END_DATA_BLOCK

DATA_BLOCK "IEC_Timer_0_DB"   // DB28
{ S7_Optimized_Access := 'TRUE' }
AUTHOR : Simatic
FAMILY : IEC
NAME : IEC_TMR
VERSION : 1.0
// stored: InstanceOfName IEC_TIMER
"IEC_TIMER"
BEGIN
END_DATA_BLOCK

DATA_BLOCK "Timer BUzzer AC2"   // DB30
{ S7_Optimized_Access := 'TRUE' }
AUTHOR : Simatic
FAMILY : IEC
NAME : IEC_TMR
VERSION : 1.0
// stored: InstanceOfName IEC_TIMER
"IEC_TIMER"
BEGIN
END_DATA_BLOCK

DATA_BLOCK "Timer Manual Insert"   // DB31
{ S7_Optimized_Access := 'TRUE' }
AUTHOR : Simatic
FAMILY : IEC
NAME : IEC_TMR
VERSION : 1.0
// stored: InstanceOfName IEC_TIMER
"IEC_TIMER"
BEGIN
END_DATA_BLOCK

DATA_BLOCK "Timer Modu"   // DB32
{ S7_Optimized_Access := 'TRUE' }
AUTHOR : Simatic
FAMILY : IEC
NAME : IEC_TMR
VERSION : 1.0
// stored: InstanceOfName IEC_TIMER
"IEC_TIMER"
BEGIN
END_DATA_BLOCK

DATA_BLOCK "Timer Reject/error Conveyor outfeed"   // DB33
{ S7_Optimized_Access := 'TRUE' }
AUTHOR : Simatic
FAMILY : IEC
NAME : IEC_TMR
VERSION : 1.0
// stored: InstanceOfName IEC_TIMER
"IEC_TIMER"
BEGIN
END_DATA_BLOCK

DATA_BLOCK "Delay Press Slof Focke"   // DB37
{ S7_Optimized_Access := 'TRUE' }
AUTHOR : Simatic
FAMILY : IEC
NAME : IEC_TMR
VERSION : 1.0
// stored: InstanceOfName IEC_TIMER
"IEC_TIMER"
BEGIN
END_DATA_BLOCK

DATA_BLOCK "IEC_Timer_0_DB_9"   // DB38
{ S7_Optimized_Access := 'TRUE' }
AUTHOR : Simatic
FAMILY : IEC
NAME : IEC_TMR
VERSION : 1.0
// stored: InstanceOfName IEC_TIMER
"IEC_TIMER"
BEGIN
END_DATA_BLOCK

DATA_BLOCK "IEC_Timer_Stop"   // DB41
{ S7_Optimized_Access := 'TRUE' }
AUTHOR : Simatic
FAMILY : IEC
NAME : IEC_TMR
VERSION : 1.0
// stored: InstanceOfName IEC_TIMER
"IEC_TIMER"
BEGIN
END_DATA_BLOCK

DATA_BLOCK "IEC_Timer_0_DB_1"   // DB42
{ S7_Optimized_Access := 'TRUE' }
AUTHOR : Simatic
FAMILY : IEC
NAME : IEC_TMR
VERSION : 1.0
// stored: InstanceOfName IEC_TIMER
"IEC_TIMER"
BEGIN
END_DATA_BLOCK

DATA_BLOCK "IEC_Timer_0_DB_5"   // DB45
{ S7_Optimized_Access := 'TRUE' }
AUTHOR : Simatic
FAMILY : IEC
NAME : IEC_TMR
VERSION : 1.0
// stored: InstanceOfName IEC_TIMER
"IEC_TIMER"
BEGIN
END_DATA_BLOCK

DATA_BLOCK "IEC_Timer_0_DB_4"   // DB47
{ S7_Optimized_Access := 'TRUE' }
AUTHOR : Simatic
FAMILY : IEC
NAME : IEC_TMR
VERSION : 1.0
// stored: InstanceOfName IEC_TIMER
"IEC_TIMER"
BEGIN
END_DATA_BLOCK

DATA_BLOCK "Timer Off Machine"   // DB48
{ S7_Optimized_Access := 'TRUE' }
AUTHOR : Simatic
FAMILY : IEC
NAME : IEC_TMR
VERSION : 1.0
// stored: InstanceOfName IEC_TIMER
"IEC_TIMER"
BEGIN
END_DATA_BLOCK

DATA_BLOCK "Timer Slof Jamed 2"   // DB49
{ S7_Optimized_Access := 'TRUE' }
AUTHOR : Simatic
FAMILY : IEC
NAME : IEC_TMR
VERSION : 1.0
// stored: InstanceOfName IEC_TIMER
"IEC_TIMER"
BEGIN
END_DATA_BLOCK

DATA_BLOCK "Timer Reject Slof"   // DB52
{ S7_Optimized_Access := 'TRUE' }
AUTHOR : Simatic
FAMILY : IEC
NAME : IEC_TMR
VERSION : 1.0
// stored: InstanceOfName IEC_TIMER
"IEC_TIMER"
BEGIN
END_DATA_BLOCK

DATA_BLOCK "Counter Paper Ribbon Out"   // DB55
{ S7_Optimized_Access := 'TRUE' }
AUTHOR : Simatic
FAMILY : IEC
NAME : IEC_TMR
VERSION : 1.0
// stored: InstanceOfName IEC_TIMER
"IEC_TIMER"
BEGIN
END_DATA_BLOCK

DATA_BLOCK "Timer After Copi SM5"   // DB60
{ S7_Optimized_Access := 'TRUE' }
AUTHOR : Simatic
FAMILY : IEC
NAME : IEC_TMR
VERSION : 1.0
// stored: InstanceOfName IEC_TIMER
"IEC_TIMER"
BEGIN
END_DATA_BLOCK

DATA_BLOCK "Timer After Copi SM4"   // DB65
{ S7_Optimized_Access := 'TRUE' }
AUTHOR : Simatic
FAMILY : IEC
NAME : IEC_TMR
VERSION : 1.0
// stored: InstanceOfName IEC_TIMER
"IEC_TIMER"
BEGIN
END_DATA_BLOCK

DATA_BLOCK "Counter Imaje Error"   // DB67
{ S7_Optimized_Access := 'TRUE' }
AUTHOR : Simatic
FAMILY : IEC
NAME : IEC_TMR
VERSION : 1.0
// stored: InstanceOfName IEC_TIMER
"IEC_TIMER"
BEGIN
END_DATA_BLOCK

DATA_BLOCK "Hitung Sloft Jammed Infeed"   // DB68
{ S7_Optimized_Access := 'TRUE' }
AUTHOR : Simatic
FAMILY : IEC
NAME : IEC_TMR
VERSION : 1.0
// stored: InstanceOfName IEC_TIMER
"IEC_TIMER"
BEGIN
END_DATA_BLOCK

DATA_BLOCK "tTM_TimerAddRej2"   // DB69
{ S7_Optimized_Access := 'TRUE' }
AUTHOR : Simatic
FAMILY : IEC
NAME : IEC_TMR
VERSION : 1.0
// stored: InstanceOfName IEC_TIMER
"IEC_TIMER"
BEGIN
END_DATA_BLOCK

DATA_BLOCK "Counter DownStream Stop"   // DB70
{ S7_Optimized_Access := 'TRUE' }
AUTHOR : Simatic
FAMILY : IEC
NAME : IEC_TMR
VERSION : 1.0
// stored: InstanceOfName IEC_TIMER
"IEC_TIMER"
BEGIN
END_DATA_BLOCK

DATA_BLOCK "Counter RS Pneu Error"   // DB71
{ S7_Optimized_Access := 'TRUE' }
AUTHOR : Simatic
FAMILY : IEC
NAME : IEC_TMR
VERSION : 1.0
// stored: InstanceOfName IEC_TIMER
"IEC_TIMER"
BEGIN
END_DATA_BLOCK

DATA_BLOCK "Counter Imaje Open"   // DB73
{ S7_Optimized_Access := 'TRUE' }
AUTHOR : Simatic
FAMILY : IEC
NAME : IEC_TMR
VERSION : 1.0
// stored: InstanceOfName IEC_TIMER
"IEC_TIMER"
BEGIN
END_DATA_BLOCK

DATA_BLOCK "Timer After Copi SM3"   // DB74
{ S7_Optimized_Access := 'TRUE' }
AUTHOR : Simatic
FAMILY : IEC
NAME : IEC_TMR
VERSION : 1.0
// stored: InstanceOfName IEC_TIMER
"IEC_TIMER"
BEGIN
END_DATA_BLOCK

DATA_BLOCK "Timer After Copi SM2"   // DB75
{ S7_Optimized_Access := 'TRUE' }
AUTHOR : Simatic
FAMILY : IEC
NAME : IEC_TMR
VERSION : 1.0
// stored: InstanceOfName IEC_TIMER
"IEC_TIMER"
BEGIN
END_DATA_BLOCK

DATA_BLOCK "Timer After Copi SM1"   // DB76
{ S7_Optimized_Access := 'TRUE' }
AUTHOR : Simatic
FAMILY : IEC
NAME : IEC_TMR
VERSION : 1.0
// stored: InstanceOfName IEC_TIMER
"IEC_TIMER"
BEGIN
END_DATA_BLOCK

DATA_BLOCK "Time Hapus data"   // DB78
{ S7_Optimized_Access := 'TRUE' }
AUTHOR : Simatic
FAMILY : IEC
NAME : IEC_TMR
VERSION : 1.0
// stored: InstanceOfName IEC_TIMER
"IEC_TIMER"
BEGIN
END_DATA_BLOCK

DATA_BLOCK "tTM_DelayReject"   // DB79
{ S7_Optimized_Access := 'TRUE' }
AUTHOR : Simatic
FAMILY : IEC
NAME : IEC_TMR
VERSION : 1.0
// stored: InstanceOfName IEC_TIMER
"IEC_TIMER"
BEGIN
END_DATA_BLOCK

DATA_BLOCK "Counter Always Bad Read"   // DB80
{ S7_Optimized_Access := 'TRUE' }
AUTHOR : Simatic
FAMILY : IEC
NAME : CNTR
VERSION : 1.0
// stored: InstanceOfName IEC_COUNTER
"IEC_COUNTER"
BEGIN
END_DATA_BLOCK

DATA_BLOCK "Timer Reset counter Always bad Read"   // DB81
{ S7_Optimized_Access := 'TRUE' }
AUTHOR : Simatic
FAMILY : IEC
NAME : IEC_TMR
VERSION : 1.0
// stored: InstanceOfName IEC_TIMER
"IEC_TIMER"
BEGIN
END_DATA_BLOCK

DATA_BLOCK "Timer paper Or Ribbon Low"   // DB82
{ S7_Optimized_Access := 'TRUE' }
AUTHOR : Simatic
FAMILY : IEC
NAME : IEC_TMR
VERSION : 1.0
// stored: InstanceOfName IEC_TIMER
"IEC_TIMER"
BEGIN
END_DATA_BLOCK

DATA_BLOCK "tTM_TimerAddRej3"   // DB83
{ S7_Optimized_Access := 'TRUE' }
AUTHOR : Simatic
FAMILY : IEC
NAME : IEC_TMR
VERSION : 1.0
// stored: InstanceOfName IEC_TIMER
"IEC_TIMER"
BEGIN
END_DATA_BLOCK

DATA_BLOCK "Timer Stop Baca"   // DB84
{ S7_Optimized_Access := 'TRUE' }
AUTHOR : Simatic
FAMILY : IEC
NAME : IEC_TMR
VERSION : 1.0
// stored: InstanceOfName IEC_TIMER
"IEC_TIMER"
BEGIN
END_DATA_BLOCK

DATA_BLOCK "Timer Mesin Running"   // DB85
{ S7_Optimized_Access := 'TRUE' }
AUTHOR : Simatic
FAMILY : IEC
NAME : IEC_TMR
VERSION : 1.0
// stored: InstanceOfName IEC_TIMER
"IEC_TIMER"
BEGIN
END_DATA_BLOCK

DATA_BLOCK "Timer Mesin Running Baypass"   // DB86
{ S7_Optimized_Access := 'TRUE' }
AUTHOR : Simatic
FAMILY : IEC
NAME : IEC_TMR
VERSION : 1.0
// stored: InstanceOfName IEC_TIMER
"IEC_TIMER"
BEGIN
END_DATA_BLOCK

DATA_BLOCK "Timer Mesin Stop"   // DB87
{ S7_Optimized_Access := 'TRUE' }
AUTHOR : Simatic
FAMILY : IEC
NAME : IEC_TMR
VERSION : 1.0
// stored: InstanceOfName IEC_TIMER
"IEC_TIMER"
BEGIN
END_DATA_BLOCK

DATA_BLOCK "Timer Mesin error"   // DB88
{ S7_Optimized_Access := 'TRUE' }
AUTHOR : Simatic
FAMILY : IEC
NAME : IEC_TMR
VERSION : 1.0
// stored: InstanceOfName IEC_TIMER
"IEC_TIMER"
BEGIN
END_DATA_BLOCK

DATA_BLOCK "tM_Counter Always Bad Read"   // DB90
{ S7_Optimized_Access := 'TRUE' }
AUTHOR : Simatic
FAMILY : IEC
NAME : IEC_TMR
VERSION : 1.0
// stored: InstanceOfName IEC_TIMER
"IEC_TIMER"
BEGIN
END_DATA_BLOCK

DATA_BLOCK "Counter Pressure Low"   // DB91
{ S7_Optimized_Access := 'TRUE' }
AUTHOR : Simatic
FAMILY : IEC
NAME : IEC_TMR
VERSION : 1.0
// stored: InstanceOfName IEC_TIMER
"IEC_TIMER"
BEGIN
END_DATA_BLOCK

DATA_BLOCK "tTM_CounterDoorOpen"   // DB92
{ S7_Optimized_Access := 'TRUE' }
AUTHOR : Simatic
FAMILY : IEC
NAME : IEC_TMR
VERSION : 1.0
// stored: InstanceOfName IEC_TIMER
"IEC_TIMER"
BEGIN
END_DATA_BLOCK

DATA_BLOCK "tTM_TimerAddRej4"   // DB93
{ S7_Optimized_Access := 'TRUE' }
AUTHOR : Simatic
FAMILY : IEC
NAME : IEC_TMR
VERSION : 1.0
// stored: InstanceOfName IEC_TIMER
"IEC_TIMER"
BEGIN
END_DATA_BLOCK

DATA_BLOCK "tTM_TimerAddRej5"   // DB94
{ S7_Optimized_Access := 'TRUE' }
AUTHOR : Simatic
FAMILY : IEC
NAME : IEC_TMR
VERSION : 1.0
// stored: InstanceOfName IEC_TIMER
"IEC_TIMER"
BEGIN
END_DATA_BLOCK

DATA_BLOCK "tTM_TimerAddRej6"   // DB95
{ S7_Optimized_Access := 'TRUE' }
AUTHOR : Simatic
FAMILY : IEC
NAME : IEC_TMR
VERSION : 1.0
// stored: InstanceOfName IEC_TIMER
"IEC_TIMER"
BEGIN
END_DATA_BLOCK

DATA_BLOCK "tTM_TimerRS1_Adv"   // DB97
{ S7_Optimized_Access := 'TRUE' }
AUTHOR : Simatic
FAMILY : IEC
NAME : IEC_TMR
VERSION : 1.0
// stored: InstanceOfName IEC_TIMER
"IEC_TIMER"
BEGIN
END_DATA_BLOCK

DATA_BLOCK "tTM_TimerRS2_Ret"   // DB99
{ S7_Optimized_Access := 'TRUE' }
AUTHOR : Simatic
FAMILY : IEC
NAME : IEC_TMR
VERSION : 1.0
// stored: InstanceOfName IEC_TIMER
"IEC_TIMER"
BEGIN
END_DATA_BLOCK

DATA_BLOCK "tTM_ErrorReject"   // DB100
{ S7_Optimized_Access := 'TRUE' }
AUTHOR : Simatic
FAMILY : IEC
NAME : IEC_TMR
VERSION : 1.0
// stored: InstanceOfName IEC_TIMER
"IEC_TIMER"
BEGIN
END_DATA_BLOCK

DATA_BLOCK "tTM_ErrorAllRSAddReject"   // DB101
{ S7_Optimized_Access := 'TRUE' }
AUTHOR : Simatic
FAMILY : IEC
NAME : IEC_TMR
VERSION : 1.0
// stored: InstanceOfName IEC_TIMER
"IEC_TIMER"
BEGIN
END_DATA_BLOCK

DATA_BLOCK "tTM_DelayNonReject"   // DB103
{ S7_Optimized_Access := 'TRUE' }
AUTHOR : Simatic
FAMILY : IEC
NAME : IEC_TMR
VERSION : 1.0
// stored: InstanceOfName IEC_TIMER
"IEC_TIMER"
BEGIN
END_DATA_BLOCK

DATA_BLOCK "tTM_ErrorNonReject"   // DB104
{ S7_Optimized_Access := 'TRUE' }
AUTHOR : Simatic
FAMILY : IEC
NAME : IEC_TMR
VERSION : 1.0
// stored: InstanceOfName IEC_TIMER
"IEC_TIMER"
BEGIN
END_DATA_BLOCK

DATA_BLOCK "tTM_CountAddReject"   // DB105
{ S7_Optimized_Access := 'TRUE' }
AUTHOR : Simatic
FAMILY : IEC
NAME : IEC_TMR
VERSION : 1.0
// stored: InstanceOfName IEC_TIMER
"IEC_TIMER"
BEGIN
END_DATA_BLOCK

// folder: (top level)

FUNCTION_BLOCK "Block Error Mode"   // FB1, LAD
{ S7_Optimized_Access := 'TRUE' }
VERSION : 0.1
   VAR_TEMP   // added for the SCL form of the ladder/FBD networks
      _w1 : Bool;
   END_VAR
BEGIN

REGION Network 1: Emergency Stop Push